// TIA Portal project "EbAndon v4_0_02" (V15) (continued)
VAR_GLOBAL   // PLC tag table "Default tag table"
   "System_Byte" AT %MB1 : Byte;
   "FirstScan" AT %M1.0 : Bool;
   "DiagStatUpdt" AT %M1.1 : Bool;
   "AlwaysTRUE" AT %M1.2 : Bool;
   "AlwaysFALSE" AT %M1.3 : Bool;
   "Clock_Byte" AT %MB0 : Byte;
   "Clock_10Hz" AT %M0.0 : Bool;
   "Clock_5Hz" AT %M0.1 : Bool;
   "Clock_2.5Hz" AT %M0.2 : Bool;
   "Clock_2Hz" AT %M0.3 : Bool;
   "Clock_1.25Hz" AT %M0.4 : Bool;
   "Clock_1Hz" AT %M0.5 : Bool;
   "Clock_0.625Hz" AT %M0.6 : Bool;
   "Clock_0.5Hz" AT %M0.7 : Bool;
   "Temp Reset" AT %M2.0 : Bool;
   "clearPartData" AT %M100.0 : Bool;
   "setDefaultPresets" AT %M100.1 : Bool;
   "hardInitReq" AT %M100.2 : Bool;
   "dbg" AT %M500.0 : Bool;
   "dbgSetDefTimes" AT %M5000.0 : Bool;
   "Copy PN Codes Into Recipes" AT %M10.0 : Bool;
   "Load Default Recipes Into Stations" AT %M10.1 : Bool;
   "Load Default Wip Data" AT %M10.2 : Bool;
END_VAR

VAR_GLOBAL   // PLC tag table "VOLVO 16 01"
   "VOLVO 16 01 IO" AT %QD1000 : DWord;
   "VOLVO 16 01 KP8 In" AT %ID0 : DWord;
   "VOLVO 16 01 KP8 Out" AT %QD0 : DWord;
END_VAR

VAR_GLOBAL   // PLC tag table "VOLVO 16 02"
   "VOLVO 16 02 IO" AT %QD1004 : DWord;
   "VOLVO 16 02 KP8 In" AT %ID4 : DWord;
   "VOLVO 16 02 KP8 Out" AT %QD4 : DWord;
END_VAR

VAR_GLOBAL   // PLC tag table "VOLVO 16 03"
   "VOLVO 16 03 IO" AT %QD1008 : DWord;
   "VOLVO 16 03 KP8 In" AT %ID8 : DWord;
   "VOLVO 16 03 KP8 Out" AT %QD8 : DWord;
END_VAR

VAR_GLOBAL   // PLC tag table "VOLVO 16 04"
   "VOLVO 16 04 IO" AT %QD1012 : DWord;
   "VOLVO 16 04 KP8 In" AT %ID12 : DWord;
   "VOLVO 16 04 KP8 Out" AT %QD12 : DWord;
END_VAR

VAR_GLOBAL   // PLC tag table "VOLVO 16 05"
   "VOLVO 16 05 IO" AT %QD1016 : DWord;
   "VOLVO 16 05 KP8 In" AT %ID16 : DWord;
   "VOLVO 16 05 KP8 Out" AT %QD16 : DWord;
END_VAR

VAR_GLOBAL   // PLC tag table "VOLVO 16 06"
   "VOLVO 16 06 IO" AT %QD1020 : DWord;
   "VOLVO 16 06 KP8 In" AT %ID20 : DWord;
   "VOLVO 16 06 KP8 Out" AT %QD20 : DWord;
END_VAR

VAR_GLOBAL   // PLC tag table "VOLVO 16 07"
   "VOLVO 16 07 IO" AT %QD1024 : DWord;
   "VOLVO 16 07 KP8 In" AT %ID24 : DWord;
   "VOLVO 16 07 KP8 Out" AT %QD24 : DWord;
END_VAR

VAR_GLOBAL   // PLC tag table "VOLVO 16 08"
   "VOLVO 16 08 IO" AT %QD1028 : DWord;
   "VOLVO 16 08 KP8 In" AT %ID28 : DWord;
   "VOLVO 16 08 KP8 Out" AT %QD28 : DWord;
END_VAR

VAR_GLOBAL   // PLC tag table "VOLVO 16 09"
   "VOLVO 16 09 IO" AT %QD1032 : DWord;
   "VOLVO 16 09 KP8 In" AT %ID32 : DWord;
   "VOLVO 16 09 KP8 Out" AT %QD32 : DWord;
END_VAR

VAR_GLOBAL   // PLC tag table "VOLVO 16 10"
   "VOLVO 16 10 IO" AT %QD1036 : DWord;
   "VOLVO 16 10 KP8 In" AT %ID36 : DWord;
   "VOLVO 16 10 KP8 Out" AT %QD36 : DWord;
END_VAR

VAR_GLOBAL   // PLC tag table "VOLVO 16 11"
   "VOLVO 16 11 IO" AT %QD1040 : DWord;
   "VOLVO 16 11 KP8 In" AT %ID40 : DWord;
   "VOLVO 16 11 KP8 Out" AT %QD40 : DWord;
END_VAR

VAR_GLOBAL   // PLC tag table "CHM 02"
   "CHM 02 KP8 In" AT %ID44 : DWord;
   "CHM 02 KP8 Out" AT %QD44 : DWord;
   "CHM 02 IO" AT %QD1044 : DWord;
END_VAR

VAR_GLOBAL   // PLC tag table "CHM 03"
   "CHM 03 IO" AT %QD1048 : DWord;
   "CHM 03 KP8 In" AT %ID48 : DWord;
   "CHM 03 KP8 Out" AT %QD48 : DWord;
END_VAR

VAR_GLOBAL   // PLC tag table "CHM 04"
   "CHM 04 IO" AT %QD1052 : DWord;
   "CHM 04 KP8 In" AT %ID52 : DWord;
   "CHM 04 KP8 Out" AT %QD52 : DWord;
END_VAR

VAR_GLOBAL   // PLC tag table "CHM 05"
   "CHM 05 IO" AT %QD1056 : DWord;
   "CHM 05 KP8 In" AT %ID56 : DWord;
   "CHM 05 KP8 Out" AT %QD56 : DWord;
END_VAR

VAR_GLOBAL   // PLC tag table "CDO 01"
   "CDO 01 IO" AT %QD1060 : DWord;
   "CDO 01 KP8 In" AT %ID60 : DWord;
   "CDO 01 KP8 Out" AT %QD60 : DWord;
END_VAR

VAR_GLOBAL   // PLC tag table "CDO 02"
   "CDO 02 IO" AT %QD1064 : DWord;
   "CDO 02 KP8 In" AT %ID64 : DWord;
   "CDO 02 KP8 Out" AT %QD64 : DWord;
END_VAR

VAR_GLOBAL   // PLC tag table "CDO 03"
   "CDO 03 IO" AT %QD1068 : DWord;
   "CDO 03 KP8 In" AT %ID68 : DWord;
   "CDO 03 KP8 Out" AT %QD68 : DWord;
END_VAR

VAR_GLOBAL   // PLC tag table "BFL 01"
   "BFL 01 IO" AT %QD1072 : DWord;
   "BFL 01 KP8 In" AT %ID72 : DWord;
   "BFL 01 KP8 Out" AT %QD72 : DWord;
   "Manual Operations Trigger" AT %M10.3 : Bool;
END_VAR

VAR_GLOBAL   // PLC tag table "BFL 02"
   "BFL 02 IO" AT %QD1076 : DWord;
   "BFL 02 KP8 In" AT %ID76 : DWord;
   "BFL 02 KP8 Out" AT %QD76 : DWord;
END_VAR

VAR_GLOBAL   // PLC tag table "BFL 03"
   "BFL 03 IO" AT %QD1080 : DWord;
   "BFL 03 KP8 In" AT %ID80 : DWord;
   "BFL 03 KP8 Out" AT %QD80 : DWord;
END_VAR

VAR_GLOBAL   // PLC tag table "LGS 01"
   "LGS 01 IO" AT %QD1084 : DWord;
   "LGS 01 KP8 In" AT %ID84 : DWord;
   "LGS 01 KP8 Out" AT %QD84 : DWord;
END_VAR

VAR_GLOBAL   // PLC tag table "LGS 02"
   "LGS 02 IO" AT %QD1088 : DWord;
   "LGS 02 KP8 In" AT %ID88 : DWord;
   "LGS 02 KP8 Out" AT %QD88 : DWord;
END_VAR

VAR_GLOBAL   // PLC tag table "CHM 01"
   "CHM 01 IO" AT %QD1092 : DWord;
   "CHM 01 KP8 In" AT %ID92 : DWord;
   "CHM 01 KP8 Out" AT %QD92 : DWord;
END_VAR

VAR_GLOBAL CONSTANT   // PLC tag table "Comm Diag"
   "pnioDeviceCount" : Int := 48;   // Upper limit of devices per HMI screen
   "USERDIAG_SLOTS_PER_SCREEN_UPPER_LIM" : Int := 31;   // Upper limit of slots per HMI screen
   "USERDIAG_SLOTS_PER_DEVICE_UPPER_LIM" : Int := 31;   // max number of modules per device
   "USERDIAG_DEVICES_PER_IO_SYSTEM_UPPER_LIM" : Int := 128;   // Upper limit of devices/slaves per IO-System/DP-Mastersystem
   "USERDIAG_SLOTS_PER_PLC_UPPER_LIM" : Int := 31;   // max number of local modules
   "USERDIAG_IO_SYSTEMS_UPPER_LIM" : Int := 1;   // Upper limit of IO-Systems/DP-Mastersystems
   "USERDIAG_IOSYSTEM_1" : Int := 1;   // Index for first IO-System/DP-Mastersystem
END_VAR

VAR_GLOBAL CONSTANT   // PLC tag table "Color Library"
   "BkBk" : USInt := 0;
   "BgWh" : USInt := 1;
   "FgWh" : USInt := 2;
   "FlWh" : USInt := 3;
   "BgGray" : USInt := 4;
   "FgGray" : USInt := 5;
   "FlGray" : USInt := 6;
   "BgLRd" : USInt := 7;
   "FgLRd" : USInt := 8;
   "FlLRd" : USInt := 9;
   "BgDRd" : USInt := 10;
   "FgDRd" : USInt := 11;
   "FlDrd" : USInt := 12;
   "BgLYe" : USInt := 13;
   "FgLYe" : USInt := 14;
   "FlLYe" : USInt := 15;
   "BgDYe" : USInt := 16;
   "FgDYe" : USInt := 17;
   "FlDYe" : USInt := 18;
   "BgLGr" : USInt := 19;
   "FgLGr" : USInt := 20;
   "FlLGr" : USInt := 21;
   "BgDGr" : USInt := 22;
   "FgDGr" : USInt := 23;
   "FlDGr" : USInt := 24;
   "BgLTe" : USInt := 25;
   "FgLTe" : USInt := 26;
   "FlLTe" : USInt := 27;
   "BgDTe" : USInt := 28;
   "FgDTe" : USInt := 29;
   "FlDTe" : USInt := 30;
   "BgLBl" : USInt := 31;
   "FgLBl" : USInt := 32;
   "FlLBl" : USInt := 33;
   "BgDBl" : USInt := 34;
   "FgDBl" : USInt := 35;
   "FlDBl" : USInt := 36;
   "BgLPu" : USInt := 37;
   "FgLPu" : USInt := 38;   // foreground light purple
   "FlLPu" : USInt := 39;
   "BgDPu" : USInt := 40;
   "FgDPu" : USInt := 41;
   "FlDPu" : USInt := 42;
   "disabled" : USInt := 254;
   "invisible" : USInt := 255;
   "LBlDRd" : USInt := 43;
   "DRdLBl" : USInt := 44;
   "LBlDRdFl" : USInt := 45;
   "DBlDRd" : USInt := 46;
   "DRdDBl" : USInt := 47;
   "DBlDRdFl" : USInt := 48;
END_VAR

VAR_GLOBAL CONSTANT   // PLC tag table "Station Meta Data"
   "btnCount" : Int := 7;   // one less than actual button count
   "stnCount" : Int := 38;   // one less than actual station count
   "defaultAlotted" : Real := 1800.0;
   "defaultCritical" : Real := 300.0;
   "wipCount" : Int := 49;
   "mStringLen" : Int := 40;
   "sStringLen" : Int := 20;
   "lStringLen" : Int := 60;
   "pnLibCount" : Int := 999;
END_VAR

VAR_GLOBAL   // PLC tag table "Simulation"
   "simMode" AT %M100.3 : Bool;
END_VAR

VAR_GLOBAL CONSTANT   // PLC tag table "Simulation"
   "simKP8Count" : Int := 11;
END_VAR

VAR_GLOBAL CONSTANT   // PLC tag table "Station IDs"
   "VOLVO 16 01" : Int := 0;
   "VOLVO 16 02" : Int := 1;
   "VOLVO 16 03" : Int := 2;
   "VOLVO 16 04" : Int := 3;
   "VOLVO 16 05" : Int := 4;
   "VOLVO 16 06" : Int := 5;
   "VOLVO 16 07" : Int := 6;
   "VOLVO 16 08" : Int := 7;
   "VOLVO 16 09" : Int := 8;
   "VOLVO 16 10" : Int := 9;
   "VOLVO 16 11" : Int := 10;
   "CHM 01" : Int := 11;
   "CHM 02" : Int := 12;
   "CHM 03" : Int := 13;
   "CHM 04" : Int := 14;
   "CHM 05" : Int := 15;
   "CDO 01" : Int := 16;
   "CDO 02" : Int := 17;
   "CDO 03" : Int := 18;
   "BFL 01" : Int := 19;
   "BFL 02" : Int := 20;
   "BFL 03" : Int := 21;
   "LGS 01" : Int := 22;
   "LGS 02" : Int := 23;
   "LGS 03" : Int := 24;
   "CV 01" : Int := 25;
   "CV 02" : Int := 26;
   "CV 03" : Int := 27;
   "CV 04" : Int := 28;
   "PC 01" : Int := 29;
   "PC 02" : Int := 30;
END_VAR

VAR_GLOBAL CONSTANT   // PLC tag table "LED Sign"
   "ledRowCount" : Int := 11;
END_VAR

VAR_GLOBAL CONSTANT   // PLC tag table "HMI Part Request Screen"
   "partReqHmiRowCount" : Int := 11;   // number of rows displayed on hmi
END_VAR

VAR_GLOBAL CONSTANT   // PLC tag table "HMI Settings Screen"
   "hmiSelStnCount" : Int := 11;   // labels for settings screen
END_VAR

VAR_GLOBAL CONSTANT   // PLC tag table "Part Request Data Base"
   "partReqDataRowCount" : Int := 199;
END_VAR

VAR_GLOBAL CONSTANT   // PLC tag table "HMI Select Station"
   "hmiStnCount" : Int := 4;   // number of stations using basic panel instead of kp8 (-1 for array)
   "hmiStnMenuSelScrnBtnCnt" : Int := 29;   // number of buttons on menu select screen (short and long rows use different data, -1 for array)
   "hmiStnMenuSelLblCnt" : Int := 29;   // number of labels (2 per row, short & long rows use same data, - 1 for array)
   "hmiStnPartSelScrnBtnCnt" : Int := 7;   // number of buttons on part select screen (-1 for array)
   "hmiStnTmpltBtnCnt" : Int := 1;   // number of button on the template (-1 for array)
END_VAR

VAR_GLOBAL   // PLC tag table "LGS 03"
   "LGS 03 IO" AT %QD1096 : DWord;
   "LGS 03 KP8 In" AT %ID96 : DWord;
   "LGS 03 KP8 Out" AT %QD96 : DWord;
END_VAR

VAR_GLOBAL   // PLC tag table "CV 01"
   "CV 01 IO" AT %QD1100 : DWord;
   "CV 01 KP8 In" AT %ID100 : DWord;
   "CV 01 KP8 Out" AT %QD100 : DWord;
END_VAR

VAR_GLOBAL   // PLC tag table "CV 02"
   "CV 02 IO" AT %QD1104 : DWord;
   "CV 02 KP8 In" AT %ID104 : DWord;
   "CV 02 KP8 Out" AT %QD104 : DWord;
END_VAR

VAR_GLOBAL   // PLC tag table "CV 03"
   "CV 03 IO" AT %QD1108 : DWord;
   "CV 03 KP8 In" AT %ID108 : DWord;
   "CV 03 KP8 Out" AT %QD108 : DWord;
END_VAR

VAR_GLOBAL   // PLC tag table "CV 04"
   "CV 04 IO" AT %QD1112 : DWord;
   "CV 04 KP8 In" AT %ID112 : DWord;
   "CV 04 KP8 Out" AT %QD112 : DWord;
END_VAR

VAR_GLOBAL   // PLC tag table "PC 01"
   "PC 01 IO" AT %QD1116 : DWord;
   "PC 01 KP8 In" AT %ID116 : DWord;
   "PC 01 KP8 Out" AT %QD116 : DWord;
END_VAR

VAR_GLOBAL   // PLC tag table "PC 02"
   "PC 02 IO" AT %QD1120 : DWord;
   "PC 02 KP8 In" AT %ID120 : DWord;
   "PC 02 KP8 Out" AT %QD120 : DWord;
END_VAR

VAR_GLOBAL CONSTANT   // PLC tag table "States"
   "requested" : Int := 10;
   "ordered" : Int := 20;
   "requestedCrit" : Int := 11;
   "requestedExp" : Int := 12;
   "acknowledged" : Int := 30;
   "reset" : Int := 99;
   "idle" : Int := 01;
   "orderedCrit" : Int := 21;
   "acknowledgedCrit" : Int := 31;
   "orderedExp" : Int := 22;
   "acknowledgedExp" : Int := 32;
   "tCritical" : Real := 5.0;
   "tAllotted" : Real := 10.0;
END_VAR

TYPE "Runtime Data"
   STRUCT
      asReal : Real;
      elapsed : LReal;
      mem : LReal;
   END_STRUCT;
END_TYPE

TYPE "Recipe: PN Code"
VERSION : 0.1
   STRUCT
      wipBtn : Array[0.."wipCount", 0.."btnCount"] of DInt;
   END_STRUCT;
END_TYPE

TYPE "Recipe: PN Codes"
VERSION : 0.1
   STRUCT
      stn : Array[0.."stnCount"] of "Recipe: PN Code";
   END_STRUCT;
   // stn[0].wipBtn[0,0] := 1000;
   // stn[0].wipBtn[0,1] := 1000;
   // stn[0].wipBtn[0,2] := 1000;
   // stn[0].wipBtn[0,3] := 173000;
   // stn[0].wipBtn[0,4] := 1000;
   // stn[0].wipBtn[0,5] := 1000;
   // stn[0].wipBtn[0,6] := 1000;
   // stn[0].wipBtn[0,7] := 169000;
   // stn[0].wipBtn[1,0] := 1000;
   // stn[0].wipBtn[1,1] := 1000;
   // stn[0].wipBtn[1,2] := 1000;
   // stn[0].wipBtn[1,3] := 1000;
   // stn[0].wipBtn[1,4] := 1000;
   // stn[0].wipBtn[1,5] := 1000;
   // stn[0].wipBtn[1,6] := 1000;
   // stn[0].wipBtn[1,7] := 1000;
   // stn[0].wipBtn[2,0] := 1000;
   // stn[0].wipBtn[2,1] := 1000;
   // stn[0].wipBtn[2,2] := 1000;
   // stn[0].wipBtn[2,3] := 1000;
   // stn[0].wipBtn[2,4] := 1000;
   // stn[0].wipBtn[2,5] := 1000;
   // stn[0].wipBtn[2,6] := 1000;
   // stn[0].wipBtn[2,7] := 1000;
   // stn[0].wipBtn[3,0] := 1000;
   // stn[0].wipBtn[3,1] := 1000;
   // stn[0].wipBtn[3,2] := 1000;
   // stn[0].wipBtn[3,3] := 1000;
   // stn[0].wipBtn[3,4] := 1000;
   // stn[0].wipBtn[3,5] := 1000;
   // stn[0].wipBtn[3,6] := 1000;
   // stn[0].wipBtn[3,7] := 1000;
   // stn[0].wipBtn[4,0] := 1000;
   // stn[0].wipBtn[4,1] := 1000;
   // stn[0].wipBtn[4,2] := 1000;
   // stn[0].wipBtn[4,3] := 1000;
   // stn[0].wipBtn[4,4] := 1000;
   // stn[0].wipBtn[4,5] := 1000;
   // stn[0].wipBtn[4,6] := 1000;
   // stn[0].wipBtn[4,7] := 1000;
   // stn[0].wipBtn[5,0] := 1000;
   // stn[0].wipBtn[5,1] := 1000;
   // stn[0].wipBtn[5,2] := 1000;
   // stn[0].wipBtn[5,3] := 1000;
   // stn[0].wipBtn[5,4] := 1000;
   // stn[0].wipBtn[5,5] := 1000;
   // stn[0].wipBtn[5,6] := 1000;
   // stn[0].wipBtn[5,7] := 1000;
   // stn[0].wipBtn[6,0] := 1000;
   // stn[0].wipBtn[6,1] := 1000;
   // stn[0].wipBtn[6,2] := 1000;
   // stn[0].wipBtn[6,3] := 1000;
   // stn[0].wipBtn[6,4] := 1000;
   // stn[0].wipBtn[6,5] := 1000;
   // stn[0].wipBtn[6,6] := 1000;
   // stn[0].wipBtn[6,7] := 1000;
   // stn[0].wipBtn[7,0] := 1000;
   // stn[0].wipBtn[7,1] := 1000;
   // stn[0].wipBtn[7,2] := 1000;
   // stn[0].wipBtn[7,3] := 1000;
   // stn[0].wipBtn[7,4] := 1000;
   // stn[0].wipBtn[7,5] := 1000;
   // stn[0].wipBtn[7,6] := 1000;
   // stn[0].wipBtn[7,7] := 1000;
   // stn[0].wipBtn[8,0] := 1000;
   // stn[0].wipBtn[8,1] := 1000;
   // stn[0].wipBtn[8,2] := 1000;
   // stn[0].wipBtn[8,3] := 1000;
   // stn[0].wipBtn[8,4] := 1000;
   // stn[0].wipBtn[8,5] := 1000;
   // stn[0].wipBtn[8,6] := 1000;
   // stn[0].wipBtn[8,7] := 1000;
   // stn[0].wipBtn[9,0] := 1000;
   // stn[0].wipBtn[9,1] := 1000;
   // stn[0].wipBtn[9,2] := 1000;
   // stn[0].wipBtn[9,3] := 1000;
   // stn[0].wipBtn[9,4] := 1000;
   // stn[0].wipBtn[9,5] := 1000;
   // stn[0].wipBtn[9,6] := 1000;
   // stn[0].wipBtn[9,7] := 1000;
   // stn[0].wipBtn[10,0] := 1000;
   // stn[0].wipBtn[10,1] := 1000;
   // stn[0].wipBtn[10,2] := 1000;
   // stn[0].wipBtn[10,3] := 1000;
   // stn[0].wipBtn[10,4] := 1000;
   // stn[0].wipBtn[10,5] := 1000;
   // stn[0].wipBtn[10,6] := 1000;
   // stn[0].wipBtn[10,7] := 1000;
   // stn[0].wipBtn[11,0] := 1000;
   // stn[0].wipBtn[11,1] := 1000;
   // stn[0].wipBtn[11,2] := 1000;
   // stn[0].wipBtn[11,3] := 1000;
   // stn[0].wipBtn[11,4] := 1000;
   // stn[0].wipBtn[11,5] := 1000;
   // stn[0].wipBtn[11,6] := 1000;
   // stn[0].wipBtn[11,7] := 1000;
   // stn[0].wipBtn[12,0] := 1000;
   // stn[0].wipBtn[12,1] := 1000;
   // stn[0].wipBtn[12,2] := 1000;
   // stn[0].wipBtn[12,3] := 1000;
   // stn[0].wipBtn[12,4] := 1000;
   // stn[0].wipBtn[12,5] := 1000;
   // stn[0].wipBtn[12,6] := 1000;
   // stn[0].wipBtn[12,7] := 1000;
   // stn[0].wipBtn[13,0] := 1000;
   // stn[0].wipBtn[13,1] := 1000;
   // stn[0].wipBtn[13,2] := 1000;
   // stn[0].wipBtn[13,3] := 1000;
   // stn[0].wipBtn[13,4] := 1000;
   // stn[0].wipBtn[13,5] := 1000;
   // stn[0].wipBtn[13,6] := 1000;
   // stn[0].wipBtn[13,7] := 1000;
   // stn[0].wipBtn[14,0] := 1000;
   // stn[0].wipBtn[14,1] := 1000;
   // stn[0].wipBtn[14,2] := 1000;
   // stn[0].wipBtn[14,3] := 1000;
   // stn[0].wipBtn[14,4] := 1000;
   // stn[0].wipBtn[14,5] := 1000;
   // stn[0].wipBtn[14,6] := 1000;
   // stn[0].wipBtn[14,7] := 1000;
   // stn[0].wipBtn[15,0] := 1000;
   // stn[0].wipBtn[15,1] := 1000;
   // stn[0].wipBtn[15,2] := 1000;
   // stn[0].wipBtn[15,3] := 1000;
   // stn[0].wipBtn[15,4] := 1000;
   // stn[0].wipBtn[15,5] := 1000;
   // stn[0].wipBtn[15,6] := 1000;
   // stn[0].wipBtn[15,7] := 1000;
   // stn[0].wipBtn[16,0] := 1000;
   // stn[0].wipBtn[16,1] := 1000;
   // stn[0].wipBtn[16,2] := 1000;
   // stn[0].wipBtn[16,3] := 1000;
   // stn[0].wipBtn[16,4] := 1000;
   // stn[0].wipBtn[16,5] := 1000;
   // stn[0].wipBtn[16,6] := 1000;
   // stn[0].wipBtn[16,7] := 1000;
   // stn[0].wipBtn[17,0] := 1000;
   // stn[0].wipBtn[17,1] := 1000;
   // stn[0].wipBtn[17,2] := 1000;
   // stn[0].wipBtn[17,3] := 1000;
   // stn[0].wipBtn[17,4] := 1000;
   // stn[0].wipBtn[17,5] := 1000;
   // stn[0].wipBtn[17,6] := 1000;
   // stn[0].wipBtn[17,7] := 1000;
   // stn[0].wipBtn[18,0] := 1000;
   // stn[0].wipBtn[18,1] := 1000;
   // stn[0].wipBtn[18,2] := 1000;
   // stn[0].wipBtn[18,3] := 1000;
   // stn[0].wipBtn[18,4] := 1000;
   // stn[0].wipBtn[18,5] := 1000;
   // stn[0].wipBtn[18,6] := 1000;
   // stn[0].wipBtn[18,7] := 1000;
   // stn[0].wipBtn[19,0] := 1000;
   // stn[0].wipBtn[19,1] := 1000;
   // stn[0].wipBtn[19,2] := 1000;
   // stn[0].wipBtn[19,3] := 1000;
   // stn[0].wipBtn[19,4] := 1000;
   // stn[0].wipBtn[19,5] := 1000;
   // stn[0].wipBtn[19,6] := 1000;
   // stn[0].wipBtn[19,7] := 1000;
   // stn[0].wipBtn[20,0] := 1000;
   // stn[0].wipBtn[20,1] := 1000;
   // stn[0].wipBtn[20,2] := 1000;
   // stn[0].wipBtn[20,3] := 1000;
   // stn[0].wipBtn[20,4] := 1000;
   // stn[0].wipBtn[20,5] := 1000;
   // stn[0].wipBtn[20,6] := 1000;
   // stn[0].wipBtn[20,7] := 1000;
   // stn[0].wipBtn[21,0] := 1000;
   // stn[0].wipBtn[21,1] := 1000;
   // stn[0].wipBtn[21,2] := 1000;
   // stn[0].wipBtn[21,3] := 1000;
   // stn[0].wipBtn[21,4] := 1000;
   // stn[0].wipBtn[21,5] := 1000;
   // stn[0].wipBtn[21,6] := 1000;
   // stn[0].wipBtn[21,7] := 1000;
   // stn[0].wipBtn[22,0] := 1000;
   // stn[0].wipBtn[22,1] := 1000;
   // stn[0].wipBtn[22,2] := 1000;
   // stn[0].wipBtn[22,3] := 1000;
   // stn[0].wipBtn[22,4] := 1000;
   // stn[0].wipBtn[22,5] := 1000;
   // stn[0].wipBtn[22,6] := 1000;
   // stn[0].wipBtn[22,7] := 1000;
   // stn[0].wipBtn[23,0] := 1000;
   // stn[0].wipBtn[23,1] := 1000;
   // stn[0].wipBtn[23,2] := 1000;
   // stn[0].wipBtn[23,3] := 1000;
   // stn[0].wipBtn[23,4] := 1000;
   // stn[0].wipBtn[23,5] := 1000;
   // stn[0].wipBtn[23,6] := 1000;
   // stn[0].wipBtn[23,7] := 1000;
   // stn[0].wipBtn[24,0] := 1000;
   // stn[0].wipBtn[24,1] := 1000;
   // stn[0].wipBtn[24,2] := 1000;
   // stn[0].wipBtn[24,3] := 1000;
   // stn[0].wipBtn[24,4] := 1000;
   // stn[0].wipBtn[24,5] := 1000;
   // stn[0].wipBtn[24,6] := 1000;
   // stn[0].wipBtn[24,7] := 1000;
   // stn[0].wipBtn[25,0] := 1000;
   // stn[0].wipBtn[25,1] := 1000;
   // stn[0].wipBtn[25,2] := 1000;
   // stn[0].wipBtn[25,3] := 1000;
   // stn[0].wipBtn[25,4] := 1000;
   // stn[0].wipBtn[25,5] := 1000;
   // stn[0].wipBtn[25,6] := 1000;
   // stn[0].wipBtn[25,7] := 1000;
   // stn[0].wipBtn[26,0] := 1000;
   // stn[0].wipBtn[26,1] := 1000;
   // stn[0].wipBtn[26,2] := 1000;
   // stn[0].wipBtn[26,3] := 1000;
   // stn[0].wipBtn[26,4] := 1000;
   // stn[0].wipBtn[26,5] := 1000;
   // stn[0].wipBtn[26,6] := 1000;
   // stn[0].wipBtn[26,7] := 1000;
   // stn[0].wipBtn[27,0] := 1000;
   // stn[0].wipBtn[27,1] := 1000;
   // stn[0].wipBtn[27,2] := 1000;
   // stn[0].wipBtn[27,3] := 1000;
   // stn[0].wipBtn[27,4] := 1000;
   // stn[0].wipBtn[27,5] := 1000;
   // stn[0].wipBtn[27,6] := 1000;
   // stn[0].wipBtn[27,7] := 1000;
   // stn[0].wipBtn[28,0] := 1000;
   // stn[0].wipBtn[28,1] := 1000;
   // stn[0].wipBtn[28,2] := 1000;
   // stn[0].wipBtn[28,3] := 1000;
   // stn[0].wipBtn[28,4] := 1000;
   // stn[0].wipBtn[28,5] := 1000;
   // stn[0].wipBtn[28,6] := 1000;
   // stn[0].wipBtn[28,7] := 1000;
   // stn[0].wipBtn[29,0] := 1000;
   // stn[0].wipBtn[29,1] := 1000;
   // stn[0].wipBtn[29,2] := 1000;
   // stn[0].wipBtn[29,3] := 1000;
   // stn[0].wipBtn[29,4] := 1000;
   // stn[0].wipBtn[29,5] := 1000;
   // stn[0].wipBtn[29,6] := 1000;
   // stn[0].wipBtn[29,7] := 1000;
   // stn[0].wipBtn[30,0] := 1000;
   // stn[0].wipBtn[30,1] := 1000;
   // stn[0].wipBtn[30,2] := 1000;
   // stn[0].wipBtn[30,3] := 1000;
   // stn[0].wipBtn[30,4] := 1000;
   // stn[0].wipBtn[30,5] := 1000;
   // stn[0].wipBtn[30,6] := 1000;
   // stn[0].wipBtn[30,7] := 1000;
   // stn[0].wipBtn[31,0] := 1000;
   // stn[0].wipBtn[31,1] := 1000;
   // stn[0].wipBtn[31,2] := 1000;
   // stn[0].wipBtn[31,3] := 1000;
   // stn[0].wipBtn[31,4] := 1000;
   // stn[0].wipBtn[31,5] := 1000;
   // stn[0].wipBtn[31,6] := 1000;
   // stn[0].wipBtn[31,7] := 1000;
   // stn[0].wipBtn[32,0] := 1000;
   // stn[0].wipBtn[32,1] := 1000;
   // stn[0].wipBtn[32,2] := 1000;
   // stn[0].wipBtn[32,3] := 1000;
   // stn[0].wipBtn[32,4] := 1000;
   // stn[0].wipBtn[32,5] := 1000;
   // stn[0].wipBtn[32,6] := 1000;
   // stn[0].wipBtn[32,7] := 1000;
   // stn[0].wipBtn[33,0] := 1000;
   // stn[0].wipBtn[33,1] := 1000;
   // stn[0].wipBtn[33,2] := 1000;
   // stn[0].wipBtn[33,3] := 1000;
   // stn[0].wipBtn[33,4] := 1000;
   // stn[0].wipBtn[33,5] := 1000;
   // stn[0].wipBtn[33,6] := 1000;
   // stn[0].wipBtn[33,7] := 1000;
   // stn[0].wipBtn[34,0] := 1000;
   // stn[0].wipBtn[34,1] := 1000;
   // stn[0].wipBtn[34,2] := 1000;
   // stn[0].wipBtn[34,3] := 1000;
   // stn[0].wipBtn[34,4] := 1000;
   // stn[0].wipBtn[34,5] := 1000;
   // stn[0].wipBtn[34,6] := 1000;
   // stn[0].wipBtn[34,7] := 1000;
   // stn[0].wipBtn[35,0] := 1000;
   // stn[0].wipBtn[35,1] := 1000;
   // stn[0].wipBtn[35,2] := 1000;
   // stn[0].wipBtn[35,3] := 1000;
   // stn[0].wipBtn[35,4] := 1000;
   // stn[0].wipBtn[35,5] := 1000;
   // stn[0].wipBtn[35,6] := 1000;
   // stn[0].wipBtn[35,7] := 1000;
   // stn[0].wipBtn[36,0] := 1000;
   // stn[0].wipBtn[36,1] := 1000;
   // stn[0].wipBtn[36,2] := 1000;
   // stn[0].wipBtn[36,3] := 1000;
   // stn[0].wipBtn[36,4] := 1000;
   // stn[0].wipBtn[36,5] := 1000;
   // stn[0].wipBtn[36,6] := 1000;
   // stn[0].wipBtn[36,7] := 1000;
   // stn[0].wipBtn[37,0] := 1000;
   // stn[0].wipBtn[37,1] := 1000;
   // stn[0].wipBtn[37,2] := 1000;
   // stn[0].wipBtn[37,3] := 1000;
   // stn[0].wipBtn[37,4] := 1000;
   // stn[0].wipBtn[37,5] := 1000;
   // stn[0].wipBtn[37,6] := 1000;
   // stn[0].wipBtn[37,7] := 1000;
   // stn[0].wipBtn[38,0] := 1000;
   // stn[0].wipBtn[38,1] := 1000;
   // stn[0].wipBtn[38,2] := 1000;
   // stn[0].wipBtn[38,3] := 1000;
   // stn[0].wipBtn[38,4] := 1000;
   // stn[0].wipBtn[38,5] := 1000;
   // stn[0].wipBtn[38,6] := 1000;
   // stn[0].wipBtn[38,7] := 1000;
   // stn[0].wipBtn[39,0] := 1000;
   // stn[0].wipBtn[39,1] := 1000;
   // stn[0].wipBtn[39,2] := 1000;
   // stn[0].wipBtn[39,3] := 1000;
   // stn[0].wipBtn[39,4] := 1000;
   // stn[0].wipBtn[39,5] := 1000;
   // stn[0].wipBtn[39,6] := 1000;
   // stn[0].wipBtn[39,7] := 1000;
   // stn[0].wipBtn[40,0] := 1000;
   // stn[0].wipBtn[40,1] := 1000;
   // stn[0].wipBtn[40,2] := 1000;
   // stn[0].wipBtn[40,3] := 1000;
   // stn[0].wipBtn[40,4] := 1000;
   // stn[0].wipBtn[40,5] := 1000;
   // stn[0].wipBtn[40,6] := 1000;
   // stn[0].wipBtn[40,7] := 1000;
   // stn[0].wipBtn[41,0] := 1000;
   // stn[0].wipBtn[41,1] := 1000;
   // stn[0].wipBtn[41,2] := 1000;
   // stn[0].wipBtn[41,3] := 1000;
   // stn[0].wipBtn[41,4] := 1000;
   // stn[0].wipBtn[41,5] := 1000;
   // stn[0].wipBtn[41,6] := 1000;
   // stn[0].wipBtn[41,7] := 1000;
   // stn[0].wipBtn[42,0] := 1000;
   // stn[0].wipBtn[42,1] := 1000;
   // stn[0].wipBtn[42,2] := 1000;
   // stn[0].wipBtn[42,3] := 1000;
   // stn[0].wipBtn[42,4] := 1000;
   // stn[0].wipBtn[42,5] := 1000;
   // stn[0].wipBtn[42,6] := 1000;
   // stn[0].wipBtn[42,7] := 1000;
   // stn[0].wipBtn[43,0] := 1000;
   // stn[0].wipBtn[43,1] := 1000;
   // stn[0].wipBtn[43,2] := 1000;
   // stn[0].wipBtn[43,3] := 1000;
   // stn[0].wipBtn[43,4] := 1000;
   // stn[0].wipBtn[43,5] := 1000;
   // stn[0].wipBtn[43,6] := 1000;
   // stn[0].wipBtn[43,7] := 1000;
   // stn[0].wipBtn[44,0] := 1000;
   // stn[0].wipBtn[44,1] := 1000;
   // stn[0].wipBtn[44,2] := 1000;
   // stn[0].wipBtn[44,3] := 1000;
   // stn[0].wipBtn[44,4] := 1000;
   // stn[0].wipBtn[44,5] := 1000;
   // stn[0].wipBtn[44,6] := 1000;
   // stn[0].wipBtn[44,7] := 1000;
   // stn[0].wipBtn[45,0] := 1000;
   // stn[0].wipBtn[45,1] := 1000;
   // stn[0].wipBtn[45,2] := 1000;
   // stn[0].wipBtn[45,3] := 1000;
   // stn[0].wipBtn[45,4] := 1000;
   // stn[0].wipBtn[45,5] := 1000;
   // stn[0].wipBtn[45,6] := 1000;
   // stn[0].wipBtn[45,7] := 1000;
   // stn[0].wipBtn[46,0] := 1000;
   // stn[0].wipBtn[46,1] := 1000;
   // stn[0].wipBtn[46,2] := 1000;
   // stn[0].wipBtn[46,3] := 1000;
   // stn[0].wipBtn[46,4] := 1000;
   // stn[0].wipBtn[46,5] := 1000;
   // stn[0].wipBtn[46,6] := 1000;
   // stn[0].wipBtn[46,7] := 1000;
   // stn[0].wipBtn[47,0] := 1000;
   // stn[0].wipBtn[47,1] := 1000;
   // stn[0].wipBtn[47,2] := 1000;
   // stn[0].wipBtn[47,3] := 1000;
   // stn[0].wipBtn[47,4] := 1000;
   // stn[0].wipBtn[47,5] := 1000;
   // stn[0].wipBtn[47,6] := 1000;
   // stn[0].wipBtn[47,7] := 1000;
   // stn[0].wipBtn[48,0] := 1000;
   // stn[0].wipBtn[48,1] := 1000;
   // stn[0].wipBtn[48,2] := 1000;
   // stn[0].wipBtn[48,3] := 1000;
   // stn[0].wipBtn[48,4] := 1000;
   // stn[0].wipBtn[48,5] := 1000;
   // stn[0].wipBtn[48,6] := 1000;
   // stn[0].wipBtn[48,7] := 1000;
   // stn[0].wipBtn[49,0] := 1000;
   // stn[0].wipBtn[49,1] := 1000;
   // stn[0].wipBtn[49,2] := 1000;
   // stn[0].wipBtn[49,3] := 1000;
   // stn[0].wipBtn[49,4] := 1000;
   // stn[0].wipBtn[49,5] := 1000;
   // stn[0].wipBtn[49,6] := 1000;
   // stn[0].wipBtn[49,7] := 1000;
   // stn[1].wipBtn[0,0] := 1000;
   // stn[1].wipBtn[0,1] := 1000;
   // stn[1].wipBtn[0,2] := 184000;
   // stn[1].wipBtn[0,3] := 210000;
   // stn[1].wipBtn[0,4] := 1000;
   // stn[1].wipBtn[0,5] := 1000;
   // stn[1].wipBtn[0,6] := 181000;
   // stn[1].wipBtn[0,7] := 167000;
   // stn[1].wipBtn[1,0] := 1000;
   // stn[1].wipBtn[1,1] := 1000;
   // stn[1].wipBtn[1,2] := 1000;
   // stn[1].wipBtn[1,3] := 1000;
   // stn[1].wipBtn[1,4] := 1000;
   // stn[1].wipBtn[1,5] := 1000;
   // stn[1].wipBtn[1,6] := 1000;
   // stn[1].wipBtn[1,7] := 1000;
   // stn[1].wipBtn[2,0] := 1000;
   // stn[1].wipBtn[2,1] := 1000;
   // stn[1].wipBtn[2,2] := 1000;
   // stn[1].wipBtn[2,3] := 1000;
   // stn[1].wipBtn[2,4] := 1000;
   // stn[1].wipBtn[2,5] := 1000;
   // stn[1].wipBtn[2,6] := 1000;
   // stn[1].wipBtn[2,7] := 1000;
   // stn[1].wipBtn[3,0] := 1000;
   // stn[1].wipBtn[3,1] := 1000;
   // stn[1].wipBtn[3,2] := 1000;
   // stn[1].wipBtn[3,3] := 1000;
   // stn[1].wipBtn[3,4] := 1000;
   // stn[1].wipBtn[3,5] := 1000;
   // stn[1].wipBtn[3,6] := 1000;
   // stn[1].wipBtn[3,7] := 1000;
   // stn[1].wipBtn[4,0] := 1000;
   // stn[1].wipBtn[4,1] := 1000;
   // stn[1].wipBtn[4,2] := 1000;
   // stn[1].wipBtn[4,3] := 1000;
   // stn[1].wipBtn[4,4] := 1000;
   // stn[1].wipBtn[4,5] := 1000;
   // stn[1].wipBtn[4,6] := 1000;
   // stn[1].wipBtn[4,7] := 1000;
   // stn[1].wipBtn[5,0] := 1000;
   // stn[1].wipBtn[5,1] := 1000;
   // stn[1].wipBtn[5,2] := 1000;
   // stn[1].wipBtn[5,3] := 1000;
   // stn[1].wipBtn[5,4] := 1000;
   // stn[1].wipBtn[5,5] := 1000;
   // stn[1].wipBtn[5,6] := 1000;
   // stn[1].wipBtn[5,7] := 1000;
   // stn[1].wipBtn[6,0] := 1000;
   // stn[1].wipBtn[6,1] := 1000;
   // stn[1].wipBtn[6,2] := 1000;
   // stn[1].wipBtn[6,3] := 1000;
   // stn[1].wipBtn[6,4] := 1000;
   // stn[1].wipBtn[6,5] := 1000;
   // stn[1].wipBtn[6,6] := 1000;
   // stn[1].wipBtn[6,7] := 1000;
   // stn[1].wipBtn[7,0] := 1000;
   // stn[1].wipBtn[7,1] := 1000;
   // stn[1].wipBtn[7,2] := 1000;
   // stn[1].wipBtn[7,3] := 1000;
   // stn[1].wipBtn[7,4] := 1000;
   // stn[1].wipBtn[7,5] := 1000;
   // stn[1].wipBtn[7,6] := 1000;
   // stn[1].wipBtn[7,7] := 1000;
   // stn[1].wipBtn[8,0] := 1000;
   // stn[1].wipBtn[8,1] := 1000;
   // stn[1].wipBtn[8,2] := 1000;
   // stn[1].wipBtn[8,3] := 1000;
   // stn[1].wipBtn[8,4] := 1000;
   // stn[1].wipBtn[8,5] := 1000;
   // stn[1].wipBtn[8,6] := 1000;
   // stn[1].wipBtn[8,7] := 1000;
   // stn[1].wipBtn[9,0] := 1000;
   // stn[1].wipBtn[9,1] := 1000;
   // stn[1].wipBtn[9,2] := 1000;
   // stn[1].wipBtn[9,3] := 1000;
   // stn[1].wipBtn[9,4] := 1000;
   // stn[1].wipBtn[9,5] := 1000;
   // stn[1].wipBtn[9,6] := 1000;
   // stn[1].wipBtn[9,7] := 1000;
   // stn[1].wipBtn[10,0] := 1000;
   // stn[1].wipBtn[10,1] := 1000;
   // stn[1].wipBtn[10,2] := 1000;
   // stn[1].wipBtn[10,3] := 1000;
   // stn[1].wipBtn[10,4] := 1000;
   // stn[1].wipBtn[10,5] := 1000;
   // stn[1].wipBtn[10,6] := 1000;
   // stn[1].wipBtn[10,7] := 1000;
   // stn[1].wipBtn[11,0] := 1000;
   // stn[1].wipBtn[11,1] := 1000;
   // stn[1].wipBtn[11,2] := 1000;
   // stn[1].wipBtn[11,3] := 1000;
   // stn[1].wipBtn[11,4] := 1000;
   // stn[1].wipBtn[11,5] := 1000;
   // stn[1].wipBtn[11,6] := 1000;
   // stn[1].wipBtn[11,7] := 1000;
   // stn[1].wipBtn[12,0] := 1000;
   // stn[1].wipBtn[12,1] := 1000;
   // stn[1].wipBtn[12,2] := 1000;
   // stn[1].wipBtn[12,3] := 1000;
   // stn[1].wipBtn[12,4] := 1000;
   // stn[1].wipBtn[12,5] := 1000;
   // stn[1].wipBtn[12,6] := 1000;
   // stn[1].wipBtn[12,7] := 1000;
   // stn[1].wipBtn[13,0] := 1000;
   // stn[1].wipBtn[13,1] := 1000;
   // stn[1].wipBtn[13,2] := 1000;
   // stn[1].wipBtn[13,3] := 1000;
   // stn[1].wipBtn[13,4] := 1000;
   // stn[1].wipBtn[13,5] := 1000;
   // stn[1].wipBtn[13,6] := 1000;
   // stn[1].wipBtn[13,7] := 1000;
   // stn[1].wipBtn[14,0] := 1000;
   // stn[1].wipBtn[14,1] := 1000;
   // stn[1].wipBtn[14,2] := 1000;
   // stn[1].wipBtn[14,3] := 1000;
   // stn[1].wipBtn[14,4] := 1000;
   // stn[1].wipBtn[14,5] := 1000;
   // stn[1].wipBtn[14,6] := 1000;
   // stn[1].wipBtn[14,7] := 1000;
   // stn[1].wipBtn[15,0] := 1000;
   // stn[1].wipBtn[15,1] := 1000;
   // stn[1].wipBtn[15,2] := 1000;
   // stn[1].wipBtn[15,3] := 1000;
   // stn[1].wipBtn[15,4] := 1000;
   // stn[1].wipBtn[15,5] := 1000;
   // stn[1].wipBtn[15,6] := 1000;
   // stn[1].wipBtn[15,7] := 1000;
   // stn[1].wipBtn[16,0] := 1000;
   // stn[1].wipBtn[16,1] := 1000;
   // stn[1].wipBtn[16,2] := 1000;
   // stn[1].wipBtn[16,3] := 1000;
   // stn[1].wipBtn[16,4] := 1000;
   // stn[1].wipBtn[16,5] := 1000;
   // stn[1].wipBtn[16,6] := 1000;
   // stn[1].wipBtn[16,7] := 1000;
   // stn[1].wipBtn[17,0] := 1000;
   // stn[1].wipBtn[17,1] := 1000;
   // stn[1].wipBtn[17,2] := 1000;
   // stn[1].wipBtn[17,3] := 1000;
   // stn[1].wipBtn[17,4] := 1000;
   // stn[1].wipBtn[17,5] := 1000;
   // stn[1].wipBtn[17,6] := 1000;
   // stn[1].wipBtn[17,7] := 1000;
   // stn[1].wipBtn[18,0] := 1000;
   // stn[1].wipBtn[18,1] := 1000;
   // stn[1].wipBtn[18,2] := 1000;
   // stn[1].wipBtn[18,3] := 1000;
   // stn[1].wipBtn[18,4] := 1000;
   // stn[1].wipBtn[18,5] := 1000;
   // stn[1].wipBtn[18,6] := 1000;
   // stn[1].wipBtn[18,7] := 1000;
   // stn[1].wipBtn[19,0] := 1000;
   // stn[1].wipBtn[19,1] := 1000;
   // stn[1].wipBtn[19,2] := 1000;
   // stn[1].wipBtn[19,3] := 1000;
   // stn[1].wipBtn[19,4] := 1000;
   // stn[1].wipBtn[19,5] := 1000;
   // stn[1].wipBtn[19,6] := 1000;
   // stn[1].wipBtn[19,7] := 1000;
   // stn[1].wipBtn[20,0] := 1000;
   // stn[1].wipBtn[20,1] := 1000;
   // stn[1].wipBtn[20,2] := 1000;
   // stn[1].wipBtn[20,3] := 1000;
   // stn[1].wipBtn[20,4] := 1000;
   // stn[1].wipBtn[20,5] := 1000;
   // stn[1].wipBtn[20,6] := 1000;
   // stn[1].wipBtn[20,7] := 1000;
   // stn[1].wipBtn[21,0] := 1000;
   // stn[1].wipBtn[21,1] := 1000;
   // stn[1].wipBtn[21,2] := 1000;
   // stn[1].wipBtn[21,3] := 1000;
   // stn[1].wipBtn[21,4] := 1000;
   // stn[1].wipBtn[21,5] := 1000;
   // stn[1].wipBtn[21,6] := 1000;
   // stn[1].wipBtn[21,7] := 1000;
   // stn[1].wipBtn[22,0] := 1000;
   // stn[1].wipBtn[22,1] := 1000;
   // stn[1].wipBtn[22,2] := 1000;
   // stn[1].wipBtn[22,3] := 1000;
   // stn[1].wipBtn[22,4] := 1000;
   // stn[1].wipBtn[22,5] := 1000;
   // stn[1].wipBtn[22,6] := 1000;
   // stn[1].wipBtn[22,7] := 1000;
   // stn[1].wipBtn[23,0] := 1000;
   // stn[1].wipBtn[23,1] := 1000;
   // stn[1].wipBtn[23,2] := 1000;
   // stn[1].wipBtn[23,3] := 1000;
   // stn[1].wipBtn[23,4] := 1000;
   // stn[1].wipBtn[23,5] := 1000;
   // stn[1].wipBtn[23,6] := 1000;
   // stn[1].wipBtn[23,7] := 1000;
   // stn[1].wipBtn[24,0] := 1000;
   // stn[1].wipBtn[24,1] := 1000;
   // stn[1].wipBtn[24,2] := 1000;
   // stn[1].wipBtn[24,3] := 1000;
   // stn[1].wipBtn[24,4] := 1000;
   // stn[1].wipBtn[24,5] := 1000;
   // stn[1].wipBtn[24,6] := 1000;
   // stn[1].wipBtn[24,7] := 1000;
   // stn[1].wipBtn[25,0] := 1000;
   // stn[1].wipBtn[25,1] := 1000;
   // stn[1].wipBtn[25,2] := 1000;
   // stn[1].wipBtn[25,3] := 1000;
   // stn[1].wipBtn[25,4] := 1000;
   // stn[1].wipBtn[25,5] := 1000;
   // stn[1].wipBtn[25,6] := 1000;
   // stn[1].wipBtn[25,7] := 1000;
   // stn[1].wipBtn[26,0] := 1000;
   // stn[1].wipBtn[26,1] := 1000;
   // stn[1].wipBtn[26,2] := 1000;
   // stn[1].wipBtn[26,3] := 1000;
   // stn[1].wipBtn[26,4] := 1000;
   // stn[1].wipBtn[26,5] := 1000;
   // stn[1].wipBtn[26,6] := 1000;
   // stn[1].wipBtn[26,7] := 1000;
   // stn[1].wipBtn[27,0] := 1000;
   // stn[1].wipBtn[27,1] := 1000;
   // stn[1].wipBtn[27,2] := 1000;
   // stn[1].wipBtn[27,3] := 1000;
   // stn[1].wipBtn[27,4] := 1000;
   // stn[1].wipBtn[27,5] := 1000;
   // stn[1].wipBtn[27,6] := 1000;
   // stn[1].wipBtn[27,7] := 1000;
   // stn[1].wipBtn[28,0] := 1000;
   // stn[1].wipBtn[28,1] := 1000;
   // stn[1].wipBtn[28,2] := 1000;
   // stn[1].wipBtn[28,3] := 1000;
   // stn[1].wipBtn[28,4] := 1000;
   // stn[1].wipBtn[28,5] := 1000;
   // stn[1].wipBtn[28,6] := 1000;
   // stn[1].wipBtn[28,7] := 1000;
   // stn[1].wipBtn[29,0] := 1000;
   // stn[1].wipBtn[29,1] := 1000;
   // stn[1].wipBtn[29,2] := 1000;